// TIA Portal project "消毒机" (V15.1)

(* hardware
DEVICE "S7-1200 station_1"  S7-1200 Station
   slot 0: "Rack_0"  S7-1200 Rack  Rack  V1.0
   slot 1: "PLC_1"  CPU 1212C DC/DC/DC  6ES7 212-1AE40-0XB0  V4.3
   slot 2: "DI 8/DQ 8x24VDC_1"  6ES7 223-1BH32-0XB0  V2.0
   slot 3: "CB 1241 (RS485)"  CB 1241 (RS485)  6ES7 241-1CH30-1XB0  V1.0
DEVICE "HMI_1"  KTP700 Basic PN
   slot 0: "HMI_1"  KTP700 Basic PN  6AV2 123-2GB03-0AX0  15.1.0.0
   slot 1: "HMI_RT_1"  KTP700 Basic PN  6AV2 123-2GB03-0AX0  15.1.0.0
   slot 5: "HMI_1.IE_CP_1"  PROFINET Interface  15.0.1.0
      slot 1: "PROFINET Interface_1"  PROFINET Interface
         slot 1: "Port_1"  Port
*)

// ===== PLC "PLC_1"  CPU 1212C DC/DC/DC =====
// protected blocks, not shown: "MB_RTU_Master_V4", "Modbus_DB", "fbRecipe"

VAR_GLOBAL   // PLC tag table "默认变量表"
   "E_Stop" AT %I0.0 : Bool;
   "Start" AT %I0.1 : Bool;
   "WepeXEnable" AT %Q0.1 : Bool;
   "CoolingWater" AT %Q0.2 : Bool;
   "AirCompressor" AT %Q0.4 : Bool;
   "Blower" AT %Q0.3 : Bool;
   "Peristalticpump" AT %Q0.0 : Bool;
   "1YV1" AT %Q1.0 : Bool;
   "1YV2" AT %Q1.1 : Bool;
   "2YV1" AT %Q1.2 : Bool;
   "2YV2" AT %Q1.3 : Bool;
   "3YV1" AT %Q1.4 : Bool;
   "3YV2" AT %Q1.5 : Bool;
   "4YV" AT %Q1.6 : Bool;
   "System_Byte" AT %MB1 : Byte;
   "FirstScan" AT %M1.0 : Bool;
   "DiagStatusUpdate" AT %M1.1 : Bool;
   "AlwaysTRUE" AT %M1.2 : Bool;
   "AlwaysFALSE" AT %M1.3 : Bool;
END_VAR

// folder: SystemDataTypeFolder

TYPE "MB_J_UDT"
VERSION : 0.1
   STRUCT
      In1 : UInt := 1;   // Modbus RTU station address:Standard addressing range (1 to 247as well as 0 for Broadcast) Extended addressing range (1 to 65535as well as 0 for Broadcast)
      In2 : USInt;   // Mode selection: Specifies the type of request (read, write or diagnostics)
      In3 : UDInt;   // Start address in the slave: Specifies the start address of the data that is accessed in the Modbus slave. The valid addresses are listed in the table of Modbus functions below.
      In4 : UInt := 1;   // Data length: Specifies the number of bits or words this instruction is to access. The valid lengths are listed in the table of Modbus functions below.
      In5 : Array[0..17] of Word;   // Data pointer: Points to the flag or DB address for the data to be written or read.
   END_STRUCT;
END_TYPE

TYPE "Unit"
   STRUCT
      Coolingwater : Bool;
      AirCompressor : Bool;
      Peristalticpump : Bool;
      WepeX_Enable : Bool;
      AYV1 : Bool;
      AYV2 : Bool;
      BYV1 : Bool;
      BYV2 : Bool;
      CYV1 : Bool;
      CYV2 : Bool;
      DYV : Bool;
      Blower : Bool;
      Runtime : Int;
      WepeX_Power : Int;
      Donebit : Int;
   END_STRUCT;
END_TYPE

TYPE "MdScn_Stus"
   STRUCT
      In1_Error : Bool;   // Flag for Modbus-RTU job DB error
      In2_Error : Bool;   // Flag for Modbus_Comm_Load Error bit
      In3_Status : Word;   // Error code for configure communication module for modbus
      In4_Error : Bool;   // Flag for Modbus_Master Error Bit
      In5_Status : Word;   // Error code for communicate as Modbus master
      In6_Error : DWord;   // Error stations for modbus communication
   END_STRUCT;
END_TYPE

TYPE "MdScn_Pr"
   STRUCT
      In1 : Port := 0;   // S7-1500/S7-1200: "HW identifier" from the device configuration
      In2 : UDInt := 9600;   // Selection of the data transmission rate
      In3 : UInt := 0;   // Selection of parity : 0 – None,1 – Odd,2 – Even
      In4 : USInt;   // Number of stop bits; 1 = 1 stop bit, 2 = 2 stop bits, 0, 3 to 255 = reserved
   END_STRUCT;
END_TYPE

// folder: (top level)

DATA_BLOCK "dbHMI"   // DB50
{ S7_Optimized_Access := 'FALSE' }
VERSION : 0.1
   VAR
      WepeX_PowerSPCom : Int;
      WepeX_PowerSP : Array[0..17] of Int;
      WepeX_ActpowerCom : Int;
      WepeX_Actpower : Array[0..17] of Int;
      WepeX_Statusword : Array[0..17] of Word;
      WepeX_Tempint : Array[0..17] of Int;
      ModbusAI : Array[0..7] of Word;
      Mode : Bool;
      WepeX_PowerMan : Bool;
      CoolingWaterMan : Bool;
      AirCompressorMan : Bool;
      BlowerMan : Bool;
      PeristalticpumpMan : Bool;
      "1YV1Man" : Bool;
      "1YV2Man" : Bool;
      "2YV1Man" : Bool;
      "2YV2Man" : Bool;
      "3YV1Man" : Bool;
      "3YV2Man" : Bool;
      "4YVMan" : Bool;
      WepeXP1_Statusword : Word;
      WepeXP2_Statusword : Word;
      WepeXP1通信正常 : Bool;
      WepeXP1通信不正常 : Bool;
      WepeXP1工作正常 : Bool;
      WepeXP1无反馈信号 : Bool;
      WepeXP1欠压保护 : Bool;
      WepeXP1过压保护 : Bool;
      WepeXP1过流保护 : Bool;
      WepeXP1过温保护 : Bool;
      WepeXP1磁控管故障 : Bool;
      WepeXP1浪涌保护 : Bool;
      WepeXP1高压故障 : Bool;
      WepeXP1开关管故障 : Bool;
      WepeXP1无功率信号 : Bool;
      WepeXP1Vcc保护 : Bool;
      WepeXP1通信状态 : Int;
      微波状态 : Int;
      火炬状态 : Int;
      Start : Bool;
      Stop : Bool;
      Reset : Bool;
      Running : Bool;
      气体温度 : Real;
      inUnit : "Unit";
      RecipeNum : Int;
      StepNumMan : Int;
      StepNumAuto : Int;
      StepNumCom : Int;
      Editor : Bool;
      Save : Bool;
      ActRcpUnit : "Unit";
      OutUnit : "Unit";
      Error : Word;
   END_VAR
BEGIN
END_DATA_BLOCK

DATA_BLOCK "dbRecipeData"   // DB51
{ S7_Optimized_Access := 'TRUE' }
VERSION : 0.1
   VAR RETAIN
      Unit : Array[1..32, 1..32] of "Unit";
   END_VAR
BEGIN
END_DATA_BLOCK

DATA_BLOCK "fbProcess_DB"   // DB100
{ S7_Optimized_Access := 'TRUE' }
VERSION : 0.1
// stored: InstanceOfName fbProcess
"fbProcess"
BEGIN
END_DATA_BLOCK

DATA_BLOCK "fbAI_DB"   // DB102
{ S7_Optimized_Access := 'TRUE' }
VERSION : 0.1
// stored: InstanceOfName fbAI
"fbAI"
BEGIN
END_DATA_BLOCK

FUNCTION_BLOCK "fbProcess"   // FB100, LAD
{ S7_Optimized_Access := 'TRUE' }
VERSION : 0.1
   VAR
      Running : Bool;
      "2YV1Auto" : Bool;
      "2YV2Auto" : Bool;
      "1YV1Auto" : Bool;
      "1YV2Auto" : Bool;
      CoolingWaterAuto : Bool;
      WepexPowerset : Bool;
      WepexPowerAuto : Bool;
      BlowerAuto : Bool;
      IEC_Timer_0_Instance : TON_TIME;
      IEC_Timer_0_Instance_1 : TON_TIME;
      IEC_Timer_0_Instance_2 : TON_TIME;
      fbRecipe_Instance : "fbRecipe";
      fbSequence_Instance : "fbSequence";
   END_VAR
   VAR_TEMP
      WepeX_PowerSPCom : Int;
      WepeX_PowerSP : Int;
   END_VAR
BEGIN

REGION Network 1
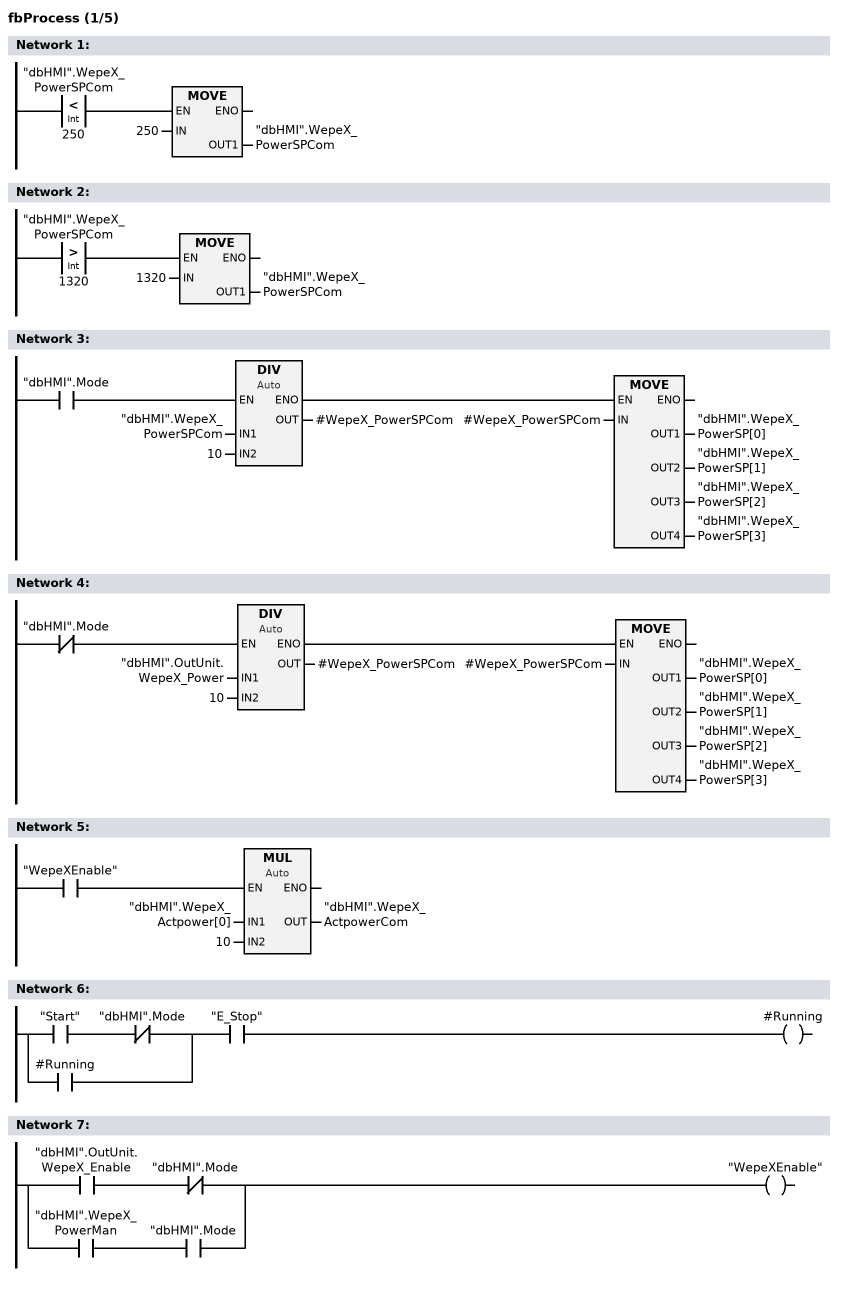
   RUNG wire#powerrail
      { S7_Templates := "SrcType := Int" } LT_Contact(in1 := "dbHMI".WepeX_PowerSPCom, in2 := 250)
      Move(in := 250, out1 => "dbHMI".WepeX_PowerSPCom)
   END_RUNG
   // the same network as SCL:
   IF "dbHMI".WepeX_PowerSPCom < 250 THEN "dbHMI".WepeX_PowerSPCom := 250; END_IF;
END_REGION

REGION Network 2
   RUNG wire#powerrail
      { S7_Templates := "SrcType := Int" } GT_Contact(in1 := "dbHMI".WepeX_PowerSPCom, in2 := 1320)
      Move(in := 1320, out1 => "dbHMI".WepeX_PowerSPCom)
   END_RUNG
   // the same network as SCL:
   IF "dbHMI".WepeX_PowerSPCom > 1320 THEN "dbHMI".WepeX_PowerSPCom := 1320; END_IF;
END_REGION

REGION Network 3
   RUNG wire#powerrail
      Contact( "dbHMI".Mode )
      Div(in1 := "dbHMI".WepeX_PowerSPCom, in2 := 10, out => #WepeX_PowerSPCom)
      Move(in := #WepeX_PowerSPCom, out1 => "dbHMI".WepeX_PowerSP[0], out2 => "dbHMI".WepeX_PowerSP[1], out3 => "dbHMI".WepeX_PowerSP[2], out4 => "dbHMI".WepeX_PowerSP[3])
   END_RUNG
   // the same network as SCL:
   IF "dbHMI".Mode THEN
       #WepeX_PowerSPCom := "dbHMI".WepeX_PowerSPCom / 10;
       "dbHMI".WepeX_PowerSP[0] := #WepeX_PowerSPCom;
       "dbHMI".WepeX_PowerSP[1] := #WepeX_PowerSPCom;
       "dbHMI".WepeX_PowerSP[2] := #WepeX_PowerSPCom;
       "dbHMI".WepeX_PowerSP[3] := #WepeX_PowerSPCom;
   END_IF;
END_REGION

REGION Network 4
   RUNG wire#powerrail
      I_Contact( "dbHMI".Mode )
      Div(in1 := "dbHMI".OutUnit.WepeX_Power, in2 := 10, out => #WepeX_PowerSPCom)
      Move(in := #WepeX_PowerSPCom, out1 => "dbHMI".WepeX_PowerSP[0], out2 => "dbHMI".WepeX_PowerSP[1], out3 => "dbHMI".WepeX_PowerSP[2], out4 => "dbHMI".WepeX_PowerSP[3])
   END_RUNG
   // the same network as SCL:
   IF NOT "dbHMI".Mode THEN
       #WepeX_PowerSPCom := "dbHMI".OutUnit.WepeX_Power / 10;
       "dbHMI".WepeX_PowerSP[0] := #WepeX_PowerSPCom;
       "dbHMI".WepeX_PowerSP[1] := #WepeX_PowerSPCom;
       "dbHMI".WepeX_PowerSP[2] := #WepeX_PowerSPCom;
       "dbHMI".WepeX_PowerSP[3] := #WepeX_PowerSPCom;
   END_IF;
END_REGION

REGION Network 5
   RUNG wire#powerrail
      Contact( "WepeXEnable" )
      Mul(in1 := "dbHMI".WepeX_Actpower[0], in2 := 10, out => "dbHMI".WepeX_ActpowerCom)
   END_RUNG
   // the same network as SCL:
   IF "WepeXEnable" THEN "dbHMI".WepeX_ActpowerCom := "dbHMI".WepeX_Actpower[0] * 10; END_IF;
END_REGION

REGION Network 6
   RUNG wire#powerrail
      Contact( "Start" )
      I_Contact( "dbHMI".Mode )
      wire#w1
      Contact( "E_Stop" )
      Coil( #Running )
   END_RUNG
   RUNG wire#powerrail
      Contact( #Running )
   END_RUNG wire#w1
   // the same network as SCL:
   #Running := (("Start" AND NOT "dbHMI".Mode) OR #Running) AND "E_Stop";
END_REGION

REGION Network 7
   RUNG wire#powerrail
      Contact( "dbHMI".OutUnit.WepeX_Enable )
      I_Contact( "dbHMI".Mode )
      wire#w1
      Coil( "WepeXEnable" )
   END_RUNG
   RUNG wire#powerrail
      Contact( "dbHMI".WepeX_PowerMan )
      Contact( "dbHMI".Mode )
   END_RUNG wire#w1
   // the same network as SCL:
   "WepeXEnable" := ("dbHMI".OutUnit.WepeX_Enable AND NOT "dbHMI".Mode) OR ("dbHMI".WepeX_PowerMan AND "dbHMI".Mode);
END_REGION

REGION Network 8
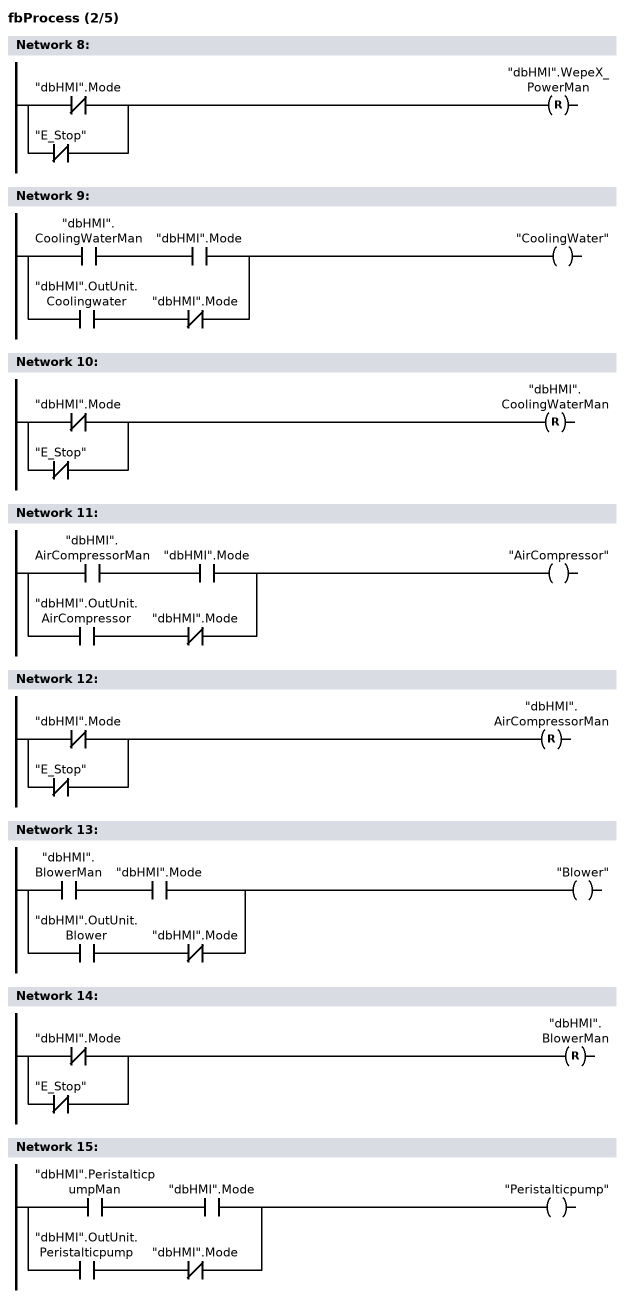
   RUNG wire#powerrail
      I_Contact( "dbHMI".Mode )
      wire#w1
      R_Coil( "dbHMI".WepeX_PowerMan )
   END_RUNG
   RUNG wire#powerrail
      I_Contact( "E_Stop" )
   END_RUNG wire#w1
   // the same network as SCL:
   IF NOT "dbHMI".Mode OR NOT "E_Stop" THEN "dbHMI".WepeX_PowerMan := FALSE; END_IF;
END_REGION

REGION Network 9
   RUNG wire#powerrail
      Contact( "dbHMI".CoolingWaterMan )
      Contact( "dbHMI".Mode )
      wire#w1
      Coil( "CoolingWater" )
   END_RUNG
   RUNG wire#powerrail
      Contact( "dbHMI".OutUnit.Coolingwater )
      I_Contact( "dbHMI".Mode )
   END_RUNG wire#w1
   // the same network as SCL:
   "CoolingWater" := ("dbHMI".CoolingWaterMan AND "dbHMI".Mode) OR ("dbHMI".OutUnit.Coolingwater AND NOT "dbHMI".Mode);
END_REGION

REGION Network 10
   RUNG wire#powerrail
      I_Contact( "dbHMI".Mode )
      wire#w1
      R_Coil( "dbHMI".CoolingWaterMan )
   END_RUNG
   RUNG wire#powerrail
      I_Contact( "E_Stop" )
   END_RUNG wire#w1
   // the same network as SCL:
   IF NOT "dbHMI".Mode OR NOT "E_Stop" THEN "dbHMI".CoolingWaterMan := FALSE; END_IF;
END_REGION

REGION Network 11
   RUNG wire#powerrail
      Contact( "dbHMI".AirCompressorMan )
      Contact( "dbHMI".Mode )
      wire#w1
      Coil( "AirCompressor" )
   END_RUNG
   RUNG wire#powerrail
      Contact( "dbHMI".OutUnit.AirCompressor )
      I_Contact( "dbHMI".Mode )
   END_RUNG wire#w1
   // the same network as SCL:
   "AirCompressor" := ("dbHMI".AirCompressorMan AND "dbHMI".Mode) OR ("dbHMI".OutUnit.AirCompressor AND NOT "dbHMI".Mode);
END_REGION

REGION Network 12
   RUNG wire#powerrail
      I_Contact( "dbHMI".Mode )
      wire#w1
      R_Coil( "dbHMI".AirCompressorMan )
   END_RUNG
   RUNG wire#powerrail
      I_Contact( "E_Stop" )
   END_RUNG wire#w1
   // the same network as SCL:
   IF NOT "dbHMI".Mode OR NOT "E_Stop" THEN "dbHMI".AirCompressorMan := FALSE; END_IF;
END_REGION

REGION Network 13
   RUNG wire#powerrail
      Contact( "dbHMI".BlowerMan )
      Contact( "dbHMI".Mode )
      wire#w1
      Coil( "Blower" )
   END_RUNG
   RUNG wire#powerrail
      Contact( "dbHMI".OutUnit.Blower )
      I_Contact( "dbHMI".Mode )
   END_RUNG wire#w1
   // the same network as SCL:
   "Blower" := ("dbHMI".BlowerMan AND "dbHMI".Mode) OR ("dbHMI".OutUnit.Blower AND NOT "dbHMI".Mode);
END_REGION

REGION Network 14
   RUNG wire#powerrail
      I_Contact( "dbHMI".Mode )
      wire#w1
      R_Coil( "dbHMI".BlowerMan )
   END_RUNG
   RUNG wire#powerrail
      I_Contact( "E_Stop" )
   END_RUNG wire#w1
   // the same network as SCL:
   IF NOT "dbHMI".Mode OR NOT "E_Stop" THEN "dbHMI".BlowerMan := FALSE; END_IF;
END_REGION

REGION Network 15
   RUNG wire#powerrail
      Contact( "dbHMI".PeristalticpumpMan )
      Contact( "dbHMI".Mode )
      wire#w1
      Coil( "Peristalticpump" )
   END_RUNG
   RUNG wire#powerrail
      Contact( "dbHMI".OutUnit.Peristalticpump )
      I_Contact( "dbHMI".Mode )
   END_RUNG wire#w1
   // the same network as SCL:
   "Peristalticpump" := ("dbHMI".PeristalticpumpMan AND "dbHMI".Mode) OR ("dbHMI".OutUnit.Peristalticpump AND NOT "dbHMI".Mode);
END_REGION

REGION Network 16
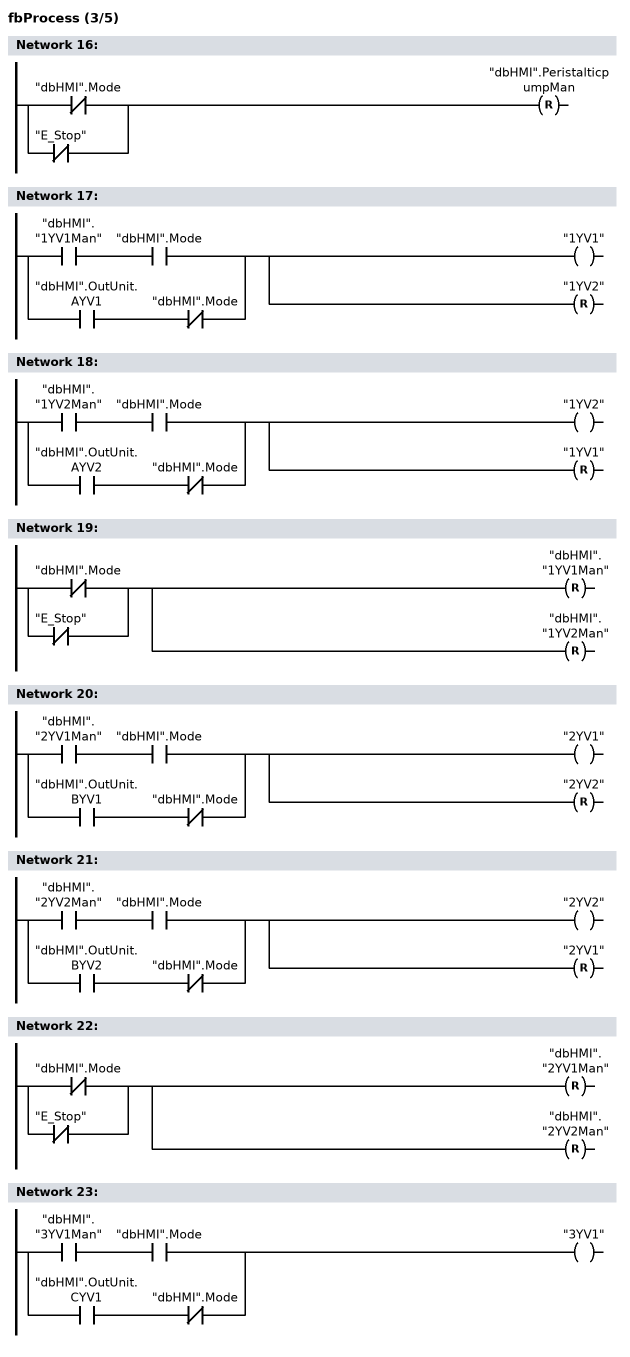
   RUNG wire#powerrail
      I_Contact( "dbHMI".Mode )
      wire#w1
      R_Coil( "dbHMI".PeristalticpumpMan )
   END_RUNG
   RUNG wire#powerrail
      I_Contact( "E_Stop" )
   END_RUNG wire#w1
   // the same network as SCL:
   IF NOT "dbHMI".Mode OR NOT "E_Stop" THEN "dbHMI".PeristalticpumpMan := FALSE; END_IF;
END_REGION

REGION Network 17
   RUNG wire#powerrail
      Contact( "dbHMI"."1YV1Man" )
      Contact( "dbHMI".Mode )
      wire#w1
      Coil( "1YV1" )
   END_RUNG
   RUNG wire#powerrail
      Contact( "dbHMI".OutUnit.AYV1 )
      I_Contact( "dbHMI".Mode )
   END_RUNG wire#w1
   RUNG wire#w1
      R_Coil( "1YV2" )
   END_RUNG
   // the same network as SCL:
   "1YV1" := ("dbHMI"."1YV1Man" AND "dbHMI".Mode) OR ("dbHMI".OutUnit.AYV1 AND NOT "dbHMI".Mode);
   IF "1YV1" THEN "1YV2" := FALSE; END_IF;
END_REGION

REGION Network 18
   RUNG wire#powerrail
      Contact( "dbHMI"."1YV2Man" )
      Contact( "dbHMI".Mode )
      wire#w1
      Coil( "1YV2" )
   END_RUNG
   RUNG wire#powerrail
      Contact( "dbHMI".OutUnit.AYV2 )
      I_Contact( "dbHMI".Mode )
   END_RUNG wire#w1
   RUNG wire#w1
      R_Coil( "1YV1" )
   END_RUNG
   // the same network as SCL:
   "1YV2" := ("dbHMI"."1YV2Man" AND "dbHMI".Mode) OR ("dbHMI".OutUnit.AYV2 AND NOT "dbHMI".Mode);
   IF "1YV2" THEN "1YV1" := FALSE; END_IF;
END_REGION

REGION Network 19
   RUNG wire#powerrail
      I_Contact( "dbHMI".Mode )
      wire#w1
      R_Coil( "dbHMI"."1YV1Man" )
   END_RUNG
   RUNG wire#powerrail
      I_Contact( "E_Stop" )
   END_RUNG wire#w1
   RUNG wire#w1
      R_Coil( "dbHMI"."1YV2Man" )
   END_RUNG
   // the same network as SCL:
   IF NOT "dbHMI".Mode OR NOT "E_Stop" THEN
       "dbHMI"."1YV1Man" := FALSE;
       "dbHMI"."1YV2Man" := FALSE;
   END_IF;
END_REGION

REGION Network 20
   RUNG wire#powerrail
      Contact( "dbHMI"."2YV1Man" )
      Contact( "dbHMI".Mode )
      wire#w1
      Coil( "2YV1" )
   END_RUNG
   RUNG wire#powerrail
      Contact( "dbHMI".OutUnit.BYV1 )
      I_Contact( "dbHMI".Mode )
   END_RUNG wire#w1
   RUNG wire#w1
      R_Coil( "2YV2" )
   END_RUNG
   // the same network as SCL:
   "2YV1" := ("dbHMI"."2YV1Man" AND "dbHMI".Mode) OR ("dbHMI".OutUnit.BYV1 AND NOT "dbHMI".Mode);
   IF "2YV1" THEN "2YV2" := FALSE; END_IF;
END_REGION

REGION Network 21
   RUNG wire#powerrail
      Contact( "dbHMI"."2YV2Man" )
      Contact( "dbHMI".Mode )
      wire#w1
      Coil( "2YV2" )
   END_RUNG
   RUNG wire#powerrail
      Contact( "dbHMI".OutUnit.BYV2 )
      I_Contact( "dbHMI".Mode )
   END_RUNG wire#w1
   RUNG wire#w1
      R_Coil( "2YV1" )
   END_RUNG
   // the same network as SCL:
   "2YV2" := ("dbHMI"."2YV2Man" AND "dbHMI".Mode) OR ("dbHMI".OutUnit.BYV2 AND NOT "dbHMI".Mode);
   IF "2YV2" THEN "2YV1" := FALSE; END_IF;
END_REGION

REGION Network 22
   RUNG wire#powerrail
      I_Contact( "dbHMI".Mode )
      wire#w1
      R_Coil( "dbHMI"."2YV1Man" )
   END_RUNG
   RUNG wire#powerrail
      I_Contact( "E_Stop" )
   END_RUNG wire#w1
   RUNG wire#w1
      R_Coil( "dbHMI"."2YV2Man" )
   END_RUNG
   // the same network as SCL:
   IF NOT "dbHMI".Mode OR NOT "E_Stop" THEN
       "dbHMI"."2YV1Man" := FALSE;
       "dbHMI"."2YV2Man" := FALSE;
   END_IF;
END_REGION

REGION Network 23
   RUNG wire#powerrail
      Contact( "dbHMI"."3YV1Man" )
      Contact( "dbHMI".Mode )
      wire#w1
      Coil( "3YV1" )
   END_RUNG
   RUNG wire#powerrail
      Contact( "dbHMI".OutUnit.CYV1 )
      I_Contact( "dbHMI".Mode )
   END_RUNG wire#w1
   // the same network as SCL:
   "3YV1" := ("dbHMI"."3YV1Man" AND "dbHMI".Mode) OR ("dbHMI".OutUnit.CYV1 AND NOT "dbHMI".Mode);
END_REGION

REGION Network 24
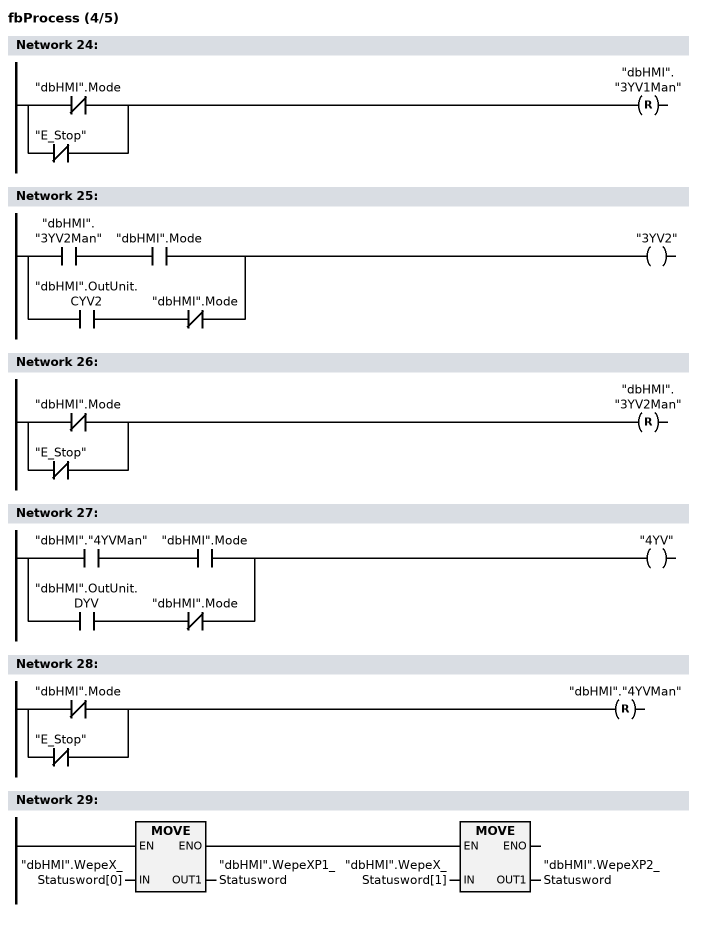
   RUNG wire#powerrail
      I_Contact( "dbHMI".Mode )
      wire#w1
      R_Coil( "dbHMI"."3YV1Man" )
   END_RUNG
   RUNG wire#powerrail
      I_Contact( "E_Stop" )
   END_RUNG wire#w1
   // the same network as SCL:
   IF NOT "dbHMI".Mode OR NOT "E_Stop" THEN "dbHMI"."3YV1Man" := FALSE; END_IF;
END_REGION

REGION Network 25
   RUNG wire#powerrail
      Contact( "dbHMI"."3YV2Man" )
      Contact( "dbHMI".Mode )
      wire#w1
      Coil( "3YV2" )
   END_RUNG
   RUNG wire#powerrail
      Contact( "dbHMI".OutUnit.CYV2 )
      I_Contact( "dbHMI".Mode )
   END_RUNG wire#w1
   // the same network as SCL:
   "3YV2" := ("dbHMI"."3YV2Man" AND "dbHMI".Mode) OR ("dbHMI".OutUnit.CYV2 AND NOT "dbHMI".Mode);
END_REGION

REGION Network 26
   RUNG wire#powerrail
      I_Contact( "dbHMI".Mode )
      wire#w1
      R_Coil( "dbHMI"."3YV2Man" )
   END_RUNG
   RUNG wire#powerrail
      I_Contact( "E_Stop" )
   END_RUNG wire#w1
   // the same network as SCL:
   IF NOT "dbHMI".Mode OR NOT "E_Stop" THEN "dbHMI"."3YV2Man" := FALSE; END_IF;
END_REGION

REGION Network 27
   RUNG wire#powerrail
      Contact( "dbHMI"."4YVMan" )
      Contact( "dbHMI".Mode )
      wire#w1
      Coil( "4YV" )
   END_RUNG
   RUNG wire#powerrail
      Contact( "dbHMI".OutUnit.DYV )
      I_Contact( "dbHMI".Mode )
   END_RUNG wire#w1
   // the same network as SCL:
   "4YV" := ("dbHMI"."4YVMan" AND "dbHMI".Mode) OR ("dbHMI".OutUnit.DYV AND NOT "dbHMI".Mode);
END_REGION

REGION Network 28
   RUNG wire#powerrail
      I_Contact( "dbHMI".Mode )
      wire#w1
      R_Coil( "dbHMI"."4YVMan" )
   END_RUNG
   RUNG wire#powerrail
      I_Contact( "E_Stop" )
   END_RUNG wire#w1
   // the same network as SCL:
   IF NOT "dbHMI".Mode OR NOT "E_Stop" THEN "dbHMI"."4YVMan" := FALSE; END_IF;
END_REGION

REGION Network 29
   RUNG wire#powerrail
      Move(in := "dbHMI".WepeX_Statusword[0], out1 => "dbHMI".WepeXP1_Statusword)
      Move(in := "dbHMI".WepeX_Statusword[1], out1 => "dbHMI".WepeXP2_Statusword)
   END_RUNG
   // the same network as SCL:
   "dbHMI".WepeXP1_Statusword := "dbHMI".WepeX_Statusword[0];
   "dbHMI".WepeXP2_Statusword := "dbHMI".WepeX_Statusword[1];
END_REGION

REGION Network 30
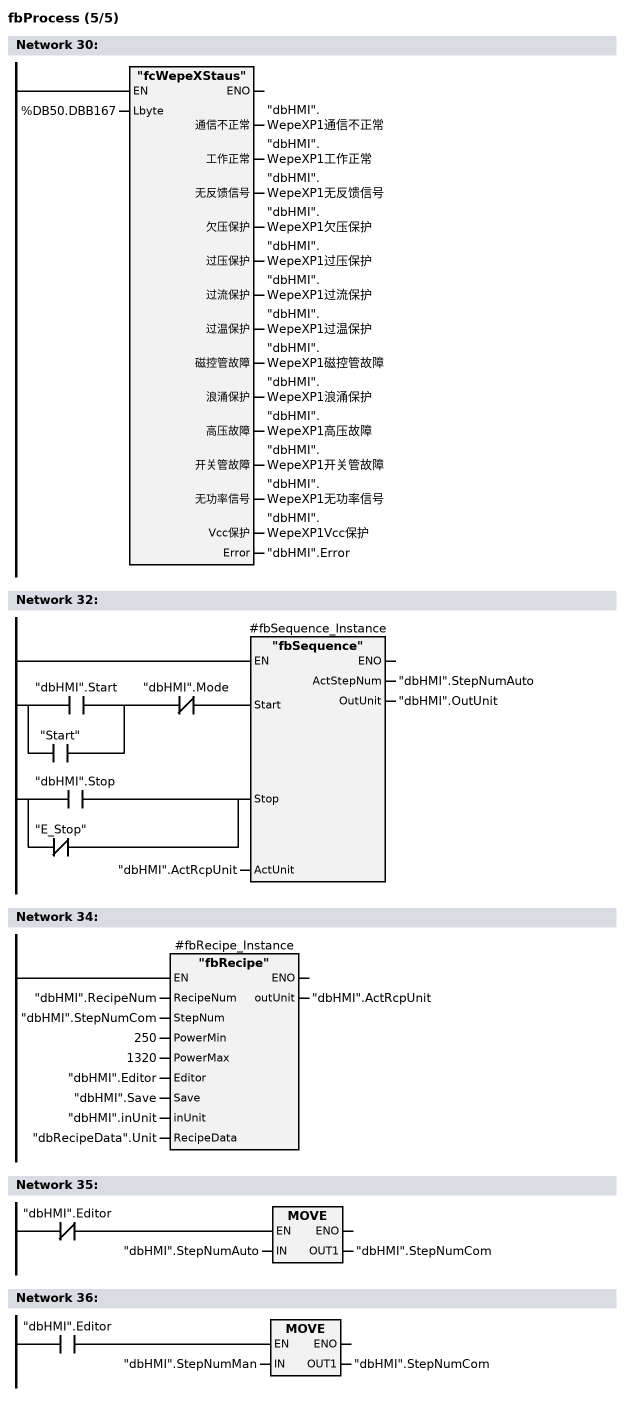
   RUNG wire#powerrail
      "fcWepeXStaus"(Lbyte := %DB50.DBB167, 通信不正常 => "dbHMI".WepeXP1通信不正常, 工作正常 => "dbHMI".WepeXP1工作正常, 无反馈信号 => "dbHMI".WepeXP1无反馈信号, 欠压保护 => "dbHMI".WepeXP1欠压保护, 过压保护 => "dbHMI".WepeXP1过压保护, 过流保护 => "dbHMI".WepeXP1过流保护, 过温保护 => "dbHMI".WepeXP1过温保护, 磁控管故障 => "dbHMI".WepeXP1磁控管故障, 浪涌保护 => "dbHMI".WepeXP1浪涌保护, 高压故障 => "dbHMI".WepeXP1高压故障, 开关管故障 => "dbHMI".WepeXP1开关管故障, 无功率信号 => "dbHMI".WepeXP1无功率信号, Vcc保护 => "dbHMI".WepeXP1Vcc保护, Error => "dbHMI".Error)
   END_RUNG
   // the same network as SCL:
   "fcWepeXStaus"(Lbyte := %DB50.DBB167,
                  通信不正常 => "dbHMI".WepeXP1通信不正常,
                  工作正常 => "dbHMI".WepeXP1工作正常,
                  无反馈信号 => "dbHMI".WepeXP1无反馈信号,
                  欠压保护 => "dbHMI".WepeXP1欠压保护,
                  过压保护 => "dbHMI".WepeXP1过压保护,
                  过流保护 => "dbHMI".WepeXP1过流保护,
                  过温保护 => "dbHMI".WepeXP1过温保护,
                  磁控管故障 => "dbHMI".WepeXP1磁控管故障,
                  浪涌保护 => "dbHMI".WepeXP1浪涌保护,
                  高压故障 => "dbHMI".WepeXP1高压故障,
                  开关管故障 => "dbHMI".WepeXP1开关管故障,
                  无功率信号 => "dbHMI".WepeXP1无功率信号,
                  Vcc保护 => "dbHMI".WepeXP1Vcc保护,
                  Error => "dbHMI".Error);
END_REGION

REGION Network 32
   RUNG wire#powerrail
      #fbSequence_Instance(Start := wire#w2, Stop := wire#w3, ActUnit := "dbHMI".ActRcpUnit, ActStepNum => "dbHMI".StepNumAuto, OutUnit => "dbHMI".OutUnit)
   END_RUNG
   RUNG wire#powerrail
      Contact( "dbHMI".Start )
      wire#w1
      I_Contact( "dbHMI".Mode )
   END_RUNG wire#w2
   RUNG wire#powerrail
      Contact( "Start" )
   END_RUNG wire#w1
   RUNG wire#powerrail
      Contact( "dbHMI".Stop )
   END_RUNG wire#w3
   RUNG wire#powerrail
      I_Contact( "E_Stop" )
   END_RUNG wire#w3
   // the same network as SCL:
   #fbSequence_Instance(Start := ("dbHMI".Start OR "Start") AND NOT "dbHMI".Mode,   // "fbSequence"
                        Stop := "dbHMI".Stop OR NOT "E_Stop",
                        ActUnit := "dbHMI".ActRcpUnit,
                        ActStepNum => "dbHMI".StepNumAuto,
                        OutUnit => "dbHMI".OutUnit);
END_REGION

REGION Network 34
   RUNG wire#powerrail
      #fbRecipe_Instance(RecipeNum := "dbHMI".RecipeNum, StepNum := "dbHMI".StepNumCom, PowerMin := 250, PowerMax := 1320, Editor := "dbHMI".Editor, Save := "dbHMI".Save, inUnit := "dbHMI".inUnit, RecipeData := "dbRecipeData".Unit, outUnit => "dbHMI".ActRcpUnit)
   END_RUNG
   // the same network as SCL:
   #fbRecipe_Instance(RecipeNum := "dbHMI".RecipeNum,   // "fbRecipe"
                      StepNum := "dbHMI".StepNumCom,
                      PowerMin := 250,
                      PowerMax := 1320,
                      Editor := "dbHMI".Editor,
                      Save := "dbHMI".Save,
                      inUnit := "dbHMI".inUnit,
                      RecipeData := "dbRecipeData".Unit,
                      outUnit => "dbHMI".ActRcpUnit);
END_REGION

REGION Network 35
   RUNG wire#powerrail
      I_Contact( "dbHMI".Editor )
      Move(in := "dbHMI".StepNumAuto, out1 => "dbHMI".StepNumCom)
   END_RUNG
   // the same network as SCL:
   IF NOT "dbHMI".Editor THEN "dbHMI".StepNumCom := "dbHMI".StepNumAuto; END_IF;
END_REGION

REGION Network 36
   RUNG wire#powerrail
      Contact( "dbHMI".Editor )
      Move(in := "dbHMI".StepNumMan, out1 => "dbHMI".StepNumCom)
   END_RUNG
   // the same network as SCL:
   IF "dbHMI".Editor THEN "dbHMI".StepNumCom := "dbHMI".StepNumMan; END_IF;
END_REGION
END_FUNCTION_BLOCK

FUNCTION_BLOCK "fbDevAI"   // FB101, LAD
{ S7_Optimized_Access := 'TRUE' }
VERSION : 0.1
   VAR_INPUT
      Norm_X_In : Word;
      Norm_X_Min : Word;
      Norm_X_Max : Word;
      Scale_X_Min : Real;
      Scale_X_Max : Real;
      Factor : Real;
      Offset : Real;
   END_VAR
   VAR_OUTPUT
      Scale_X_Out : Real;
   END_VAR
   VAR_TEMP
      temp0 : Real;
      temp1 : Real;
      temp2 : Real;
   END_VAR
BEGIN

REGION Network 1